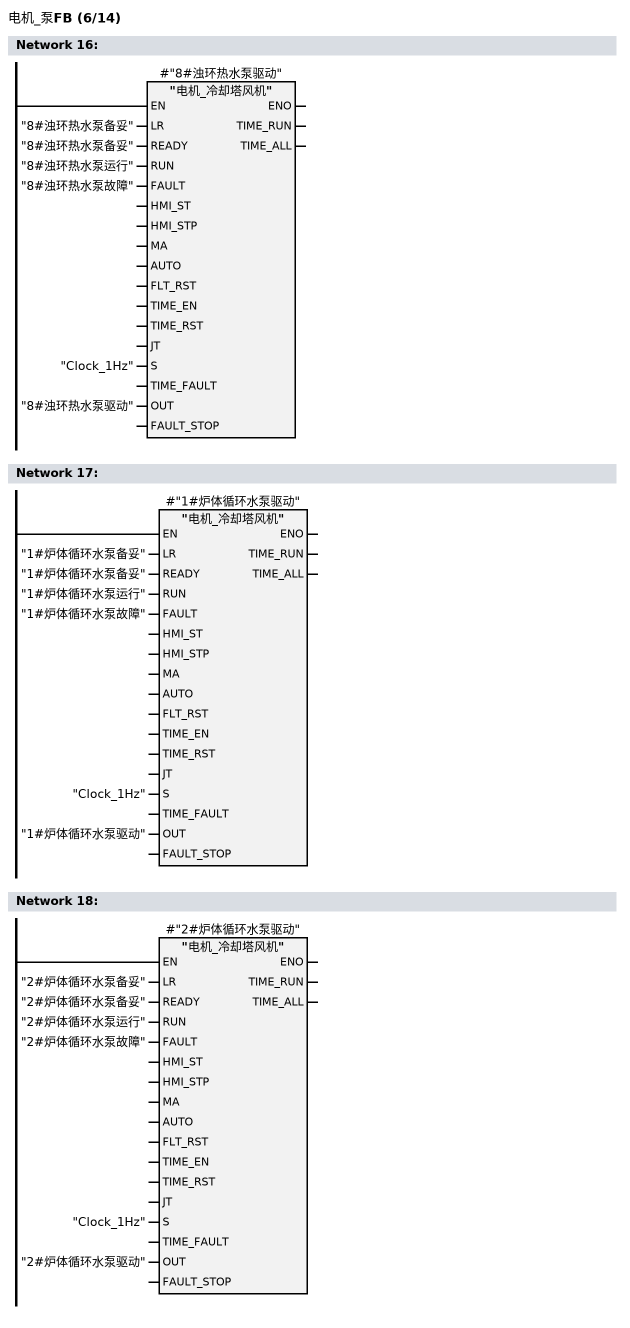
   RUNG wire#powerrail
      #"8#浊环热水泵驱动"(LR := "8#浊环热水泵备妥", READY := "8#浊环热水泵备妥", RUN := "8#浊环热水泵运行", FAULT := "8#浊环热水泵故障", HMI_ST :=, HMI_STP :=, MA :=, AUTO :=, FLT_RST :=, TIME_EN :=, TIME_RST :=, JT :=, S := "Clock_1Hz", TIME_FAULT :=, OUT := "8#浊环热水泵驱动", FAULT_STOP :=, TIME_RUN =>, TIME_ALL =>)
   END_RUNG
   // the same network as SCL:
   #"8#浊环热水泵驱动"(LR := "8#浊环热水泵备妥",   // "电机_冷却塔风机"
                READY := "8#浊环热水泵备妥",
                RUN := "8#浊环热水泵运行",
                FAULT := "8#浊环热水泵故障",
                S := "Clock_1Hz",
                OUT := "8#浊环热水泵驱动");
END_REGION

REGION Network 17
   RUNG wire#powerrail
      #"1#炉体循环水泵驱动"(LR := "1#炉体循环水泵备妥", READY := "1#炉体循环水泵备妥", RUN := "1#炉体循环水泵运行", FAULT := "1#炉体循环水泵故障", HMI_ST :=, HMI_STP :=, MA :=, AUTO :=, FLT_RST :=, TIME_EN :=, TIME_RST :=, JT :=, S := "Clock_1Hz", TIME_FAULT :=, OUT := "1#炉体循环水泵驱动", FAULT_STOP :=, TIME_RUN =>, TIME_ALL =>)
   END_RUNG
   // the same network as SCL:
   #"1#炉体循环水泵驱动"(LR := "1#炉体循环水泵备妥",   // "电机_冷却塔风机"
                 READY := "1#炉体循环水泵备妥",
                 RUN := "1#炉体循环水泵运行",
                 FAULT := "1#炉体循环水泵故障",
                 S := "Clock_1Hz",
                 OUT := "1#炉体循环水泵驱动");
END_REGION

REGION Network 18
   RUNG wire#powerrail
      #"2#炉体循环水泵驱动"(LR := "2#炉体循环水泵备妥", READY := "2#炉体循环水泵备妥", RUN := "2#炉体循环水泵运行", FAULT := "2#炉体循环水泵故障", HMI_ST :=, HMI_STP :=, MA :=, AUTO :=, FLT_RST :=, TIME_EN :=, TIME_RST :=, JT :=, S := "Clock_1Hz", TIME_FAULT :=, OUT := "2#炉体循环水泵驱动", FAULT_STOP :=, TIME_RUN =>, TIME_ALL =>)
   END_RUNG
   // the same network as SCL:
   #"2#炉体循环水泵驱动"(LR := "2#炉体循环水泵备妥",   // "电机_冷却塔风机"
                 READY := "2#炉体循环水泵备妥",
                 RUN := "2#炉体循环水泵运行",
                 FAULT := "2#炉体循环水泵故障",
                 S := "Clock_1Hz",
                 OUT := "2#炉体循环水泵驱动");
END_REGION

REGION Network 19
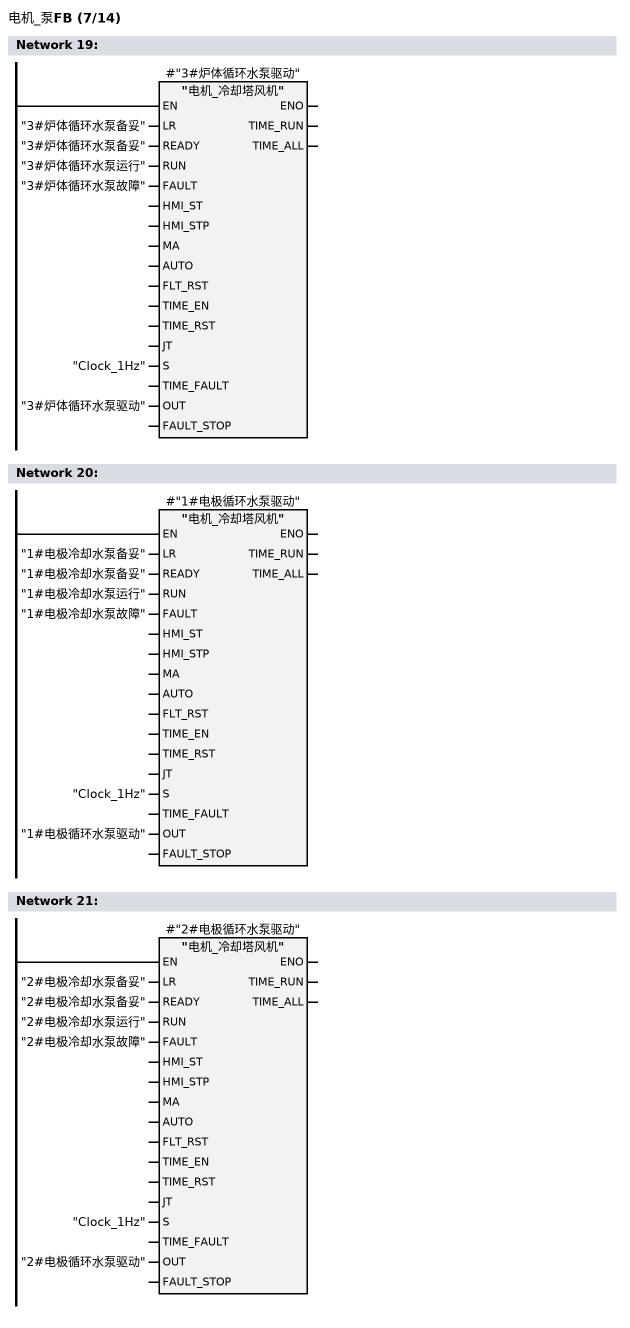
   RUNG wire#powerrail
      #"3#炉体循环水泵驱动"(LR := "3#炉体循环水泵备妥", READY := "3#炉体循环水泵备妥", RUN := "3#炉体循环水泵运行", FAULT := "3#炉体循环水泵故障", HMI_ST :=, HMI_STP :=, MA :=, AUTO :=, FLT_RST :=, TIME_EN :=, TIME_RST :=, JT :=, S := "Clock_1Hz", TIME_FAULT :=, OUT := "3#炉体循环水泵驱动", FAULT_STOP :=, TIME_RUN =>, TIME_ALL =>)
   END_RUNG
   // the same network as SCL:
   #"3#炉体循环水泵驱动"(LR := "3#炉体循环水泵备妥",   // "电机_冷却塔风机"
                 READY := "3#炉体循环水泵备妥",
                 RUN := "3#炉体循环水泵运行",
                 FAULT := "3#炉体循环水泵故障",
                 S := "Clock_1Hz",
                 OUT := "3#炉体循环水泵驱动");
END_REGION

REGION Network 20
   RUNG wire#powerrail
      #"1#电极循环水泵驱动"(LR := "1#电极冷却水泵备妥", READY := "1#电极冷却水泵备妥", RUN := "1#电极冷却水泵运行", FAULT := "1#电极冷却水泵故障", HMI_ST :=, HMI_STP :=, MA :=, AUTO :=, FLT_RST :=, TIME_EN :=, TIME_RST :=, JT :=, S := "Clock_1Hz", TIME_FAULT :=, OUT := "1#电极循环水泵驱动", FAULT_STOP :=, TIME_RUN =>, TIME_ALL =>)
   END_RUNG
   // the same network as SCL:
   #"1#电极循环水泵驱动"(LR := "1#电极冷却水泵备妥",   // "电机_冷却塔风机"
                 READY := "1#电极冷却水泵备妥",
                 RUN := "1#电极冷却水泵运行",
                 FAULT := "1#电极冷却水泵故障",
                 S := "Clock_1Hz",
                 OUT := "1#电极循环水泵驱动");
END_REGION

REGION Network 21
   RUNG wire#powerrail
      #"2#电极循环水泵驱动"(LR := "2#电极冷却水泵备妥", READY := "2#电极冷却水泵备妥", RUN := "2#电极冷却水泵运行", FAULT := "2#电极冷却水泵故障", HMI_ST :=, HMI_STP :=, MA :=, AUTO :=, FLT_RST :=, TIME_EN :=, TIME_RST :=, JT :=, S := "Clock_1Hz", TIME_FAULT :=, OUT := "2#电极循环水泵驱动", FAULT_STOP :=, TIME_RUN =>, TIME_ALL =>)
   END_RUNG
   // the same network as SCL:
   #"2#电极循环水泵驱动"(LR := "2#电极冷却水泵备妥",   // "电机_冷却塔风机"
                 READY := "2#电极冷却水泵备妥",
                 RUN := "2#电极冷却水泵运行",
                 FAULT := "2#电极冷却水泵故障",
                 S := "Clock_1Hz",
                 OUT := "2#电极循环水泵驱动");
END_REGION

REGION Network 22
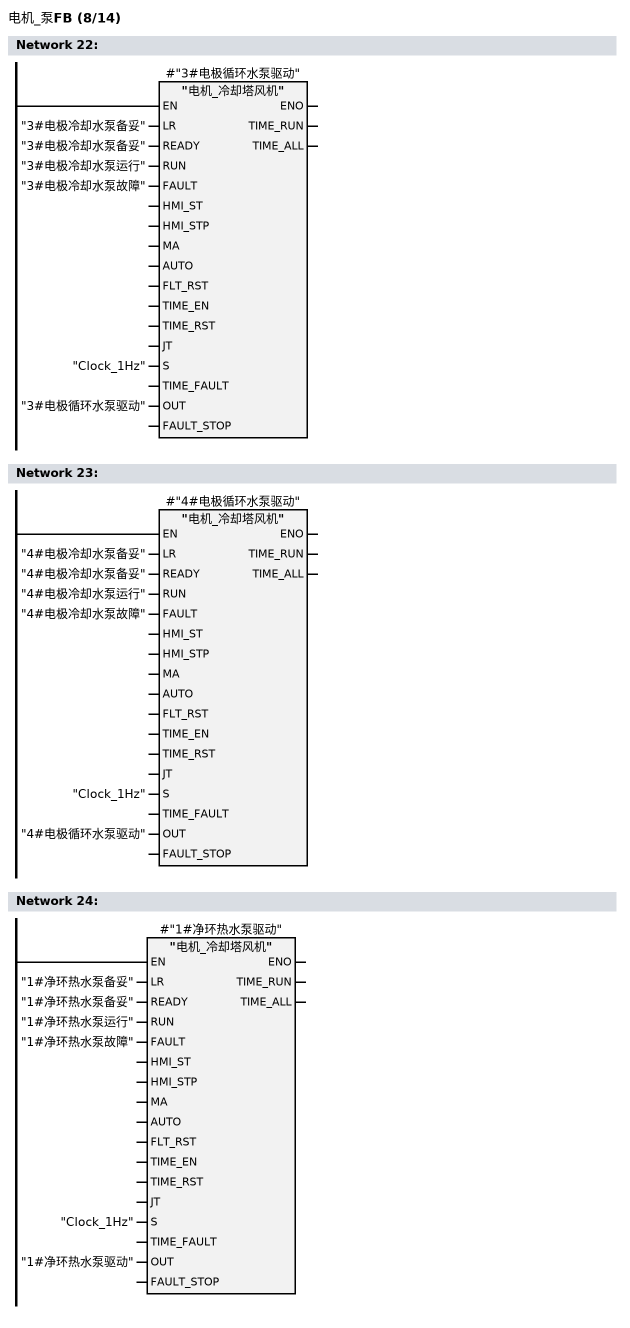
   RUNG wire#powerrail
      #"3#电极循环水泵驱动"(LR := "3#电极冷却水泵备妥", READY := "3#电极冷却水泵备妥", RUN := "3#电极冷却水泵运行", FAULT := "3#电极冷却水泵故障", HMI_ST :=, HMI_STP :=, MA :=, AUTO :=, FLT_RST :=, TIME_EN :=, TIME_RST :=, JT :=, S := "Clock_1Hz", TIME_FAULT :=, OUT := "3#电极循环水泵驱动", FAULT_STOP :=, TIME_RUN =>, TIME_ALL =>)
   END_RUNG
   // the same network as SCL:
   #"3#电极循环水泵驱动"(LR := "3#电极冷却水泵备妥",   // "电机_冷却塔风机"
                 READY := "3#电极冷却水泵备妥",
                 RUN := "3#电极冷却水泵运行",
                 FAULT := "3#电极冷却水泵故障",
                 S := "Clock_1Hz",
                 OUT := "3#电极循环水泵驱动");
END_REGION

REGION Network 23
   RUNG wire#powerrail
      #"4#电极循环水泵驱动"(LR := "4#电极冷却水泵备妥", READY := "4#电极冷却水泵备妥", RUN := "4#电极冷却水泵运行", FAULT := "4#电极冷却水泵故障", HMI_ST :=, HMI_STP :=, MA :=, AUTO :=, FLT_RST :=, TIME_EN :=, TIME_RST :=, JT :=, S := "Clock_1Hz", TIME_FAULT :=, OUT := "4#电极循环水泵驱动", FAULT_STOP :=, TIME_RUN =>, TIME_ALL =>)
   END_RUNG
   // the same network as SCL:
   #"4#电极循环水泵驱动"(LR := "4#电极冷却水泵备妥",   // "电机_冷却塔风机"
                 READY := "4#电极冷却水泵备妥",
                 RUN := "4#电极冷却水泵运行",
                 FAULT := "4#电极冷却水泵故障",
                 S := "Clock_1Hz",
                 OUT := "4#电极循环水泵驱动");
END_REGION

REGION Network 24
   RUNG wire#powerrail
      #"1#净环热水泵驱动"(LR := "1#净环热水泵备妥", READY := "1#净环热水泵备妥", RUN := "1#净环热水泵运行", FAULT := "1#净环热水泵故障", HMI_ST :=, HMI_STP :=, MA :=, AUTO :=, FLT_RST :=, TIME_EN :=, TIME_RST :=, JT :=, S := "Clock_1Hz", TIME_FAULT :=, OUT := "1#净环热水泵驱动", FAULT_STOP :=, TIME_RUN =>, TIME_ALL =>)
   END_RUNG
   // the same network as SCL:
   #"1#净环热水泵驱动"(LR := "1#净环热水泵备妥",   // "电机_冷却塔风机"
                READY := "1#净环热水泵备妥",
                RUN := "1#净环热水泵运行",
                FAULT := "1#净环热水泵故障",
                S := "Clock_1Hz",
                OUT := "1#净环热水泵驱动");
END_REGION

REGION Network 25
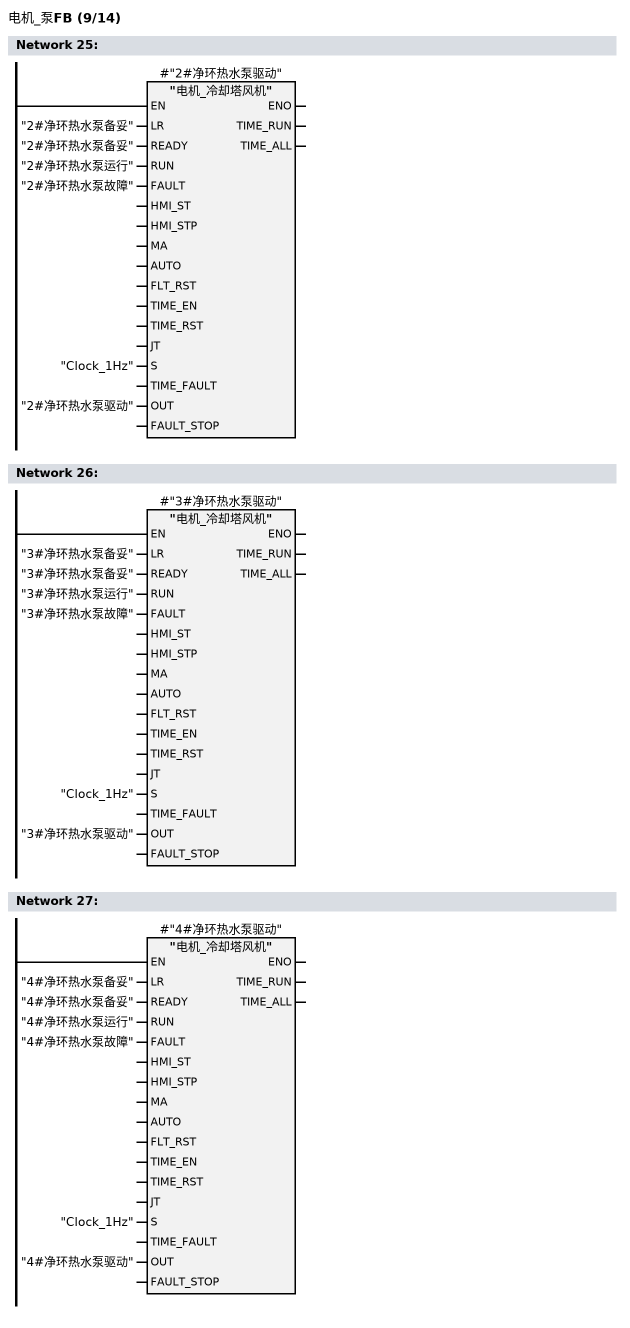
   RUNG wire#powerrail
      #"2#净环热水泵驱动"(LR := "2#净环热水泵备妥", READY := "2#净环热水泵备妥", RUN := "2#净环热水泵运行", FAULT := "2#净环热水泵故障", HMI_ST :=, HMI_STP :=, MA :=, AUTO :=, FLT_RST :=, TIME_EN :=, TIME_RST :=, JT :=, S := "Clock_1Hz", TIME_FAULT :=, OUT := "2#净环热水泵驱动", FAULT_STOP :=, TIME_RUN =>, TIME_ALL =>)
   END_RUNG
   // the same network as SCL:
   #"2#净环热水泵驱动"(LR := "2#净环热水泵备妥",   // "电机_冷却塔风机"
                READY := "2#净环热水泵备妥",
                RUN := "2#净环热水泵运行",
                FAULT := "2#净环热水泵故障",
                S := "Clock_1Hz",
                OUT := "2#净环热水泵驱动");
END_REGION

REGION Network 26
   RUNG wire#powerrail
      #"3#净环热水泵驱动"(LR := "3#净环热水泵备妥", READY := "3#净环热水泵备妥", RUN := "3#净环热水泵运行", FAULT := "3#净环热水泵故障", HMI_ST :=, HMI_STP :=, MA :=, AUTO :=, FLT_RST :=, TIME_EN :=, TIME_RST :=, JT :=, S := "Clock_1Hz", TIME_FAULT :=, OUT := "3#净环热水泵驱动", FAULT_STOP :=, TIME_RUN =>, TIME_ALL =>)
   END_RUNG
   // the same network as SCL:
   #"3#净环热水泵驱动"(LR := "3#净环热水泵备妥",   // "电机_冷却塔风机"
                READY := "3#净环热水泵备妥",
                RUN := "3#净环热水泵运行",
                FAULT := "3#净环热水泵故障",
                S := "Clock_1Hz",
                OUT := "3#净环热水泵驱动");
END_REGION

REGION Network 27
   RUNG wire#powerrail
      #"4#净环热水泵驱动"(LR := "4#净环热水泵备妥", READY := "4#净环热水泵备妥", RUN := "4#净环热水泵运行", FAULT := "4#净环热水泵故障", HMI_ST :=, HMI_STP :=, MA :=, AUTO :=, FLT_RST :=, TIME_EN :=, TIME_RST :=, JT :=, S := "Clock_1Hz", TIME_FAULT :=, OUT := "4#净环热水泵驱动", FAULT_STOP :=, TIME_RUN =>, TIME_ALL =>)
   END_RUNG
   // the same network as SCL:
   #"4#净环热水泵驱动"(LR := "4#净环热水泵备妥",   // "电机_冷却塔风机"
                READY := "4#净环热水泵备妥",
                RUN := "4#净环热水泵运行",
                FAULT := "4#净环热水泵故障",
                S := "Clock_1Hz",
                OUT := "4#净环热水泵驱动");
END_REGION

REGION Network 28
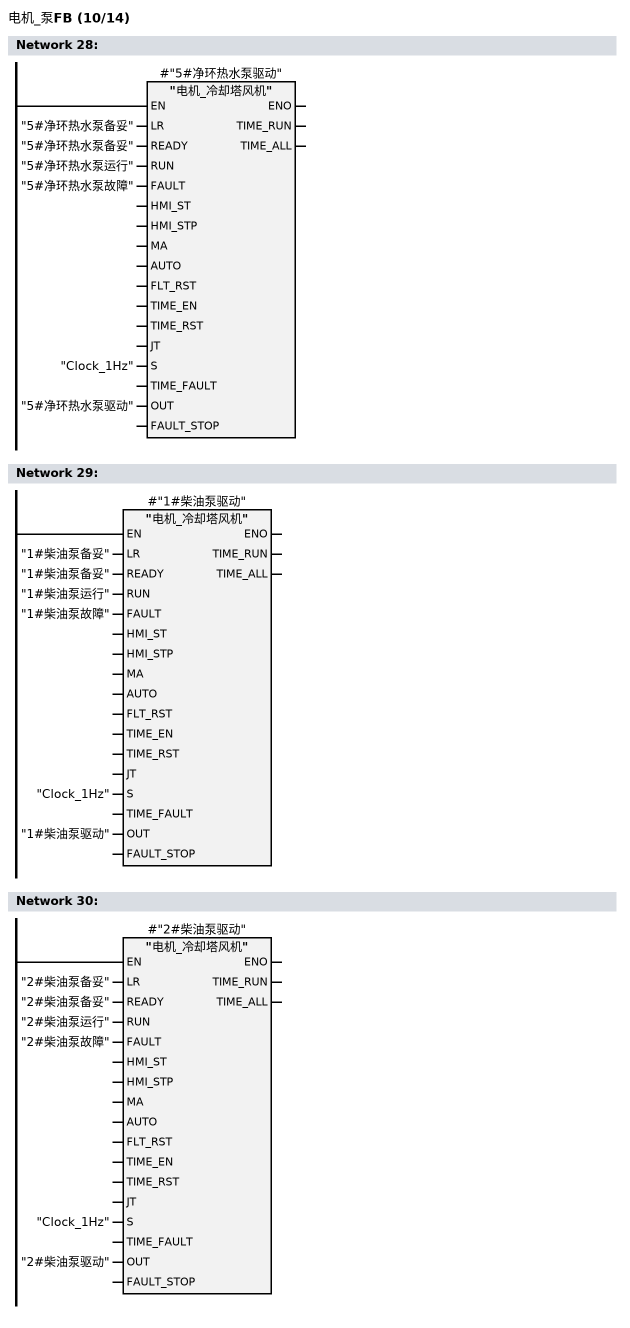
   RUNG wire#powerrail
      #"5#净环热水泵驱动"(LR := "5#净环热水泵备妥", READY := "5#净环热水泵备妥", RUN := "5#净环热水泵运行", FAULT := "5#净环热水泵故障", HMI_ST :=, HMI_STP :=, MA :=, AUTO :=, FLT_RST :=, TIME_EN :=, TIME_RST :=, JT :=, S := "Clock_1Hz", TIME_FAULT :=, OUT := "5#净环热水泵驱动", FAULT_STOP :=, TIME_RUN =>, TIME_ALL =>)
   END_RUNG
   // the same network as SCL:
   #"5#净环热水泵驱动"(LR := "5#净环热水泵备妥",   // "电机_冷却塔风机"
                READY := "5#净环热水泵备妥",
                RUN := "5#净环热水泵运行",
                FAULT := "5#净环热水泵故障",
                S := "Clock_1Hz",
                OUT := "5#净环热水泵驱动");
END_REGION

REGION Network 29
   RUNG wire#powerrail
      #"1#柴油泵驱动"(LR := "1#柴油泵备妥", READY := "1#柴油泵备妥", RUN := "1#柴油泵运行", FAULT := "1#柴油泵故障", HMI_ST :=, HMI_STP :=, MA :=, AUTO :=, FLT_RST :=, TIME_EN :=, TIME_RST :=, JT :=, S := "Clock_1Hz", TIME_FAULT :=, OUT := "1#柴油泵驱动", FAULT_STOP :=, TIME_RUN =>, TIME_ALL =>)
   END_RUNG
   // the same network as SCL:
   #"1#柴油泵驱动"(LR := "1#柴油泵备妥",   // "电机_冷却塔风机"
              READY := "1#柴油泵备妥",
              RUN := "1#柴油泵运行",
              FAULT := "1#柴油泵故障",
              S := "Clock_1Hz",
              OUT := "1#柴油泵驱动");
END_REGION

REGION Network 30
   RUNG wire#powerrail
      #"2#柴油泵驱动"(LR := "2#柴油泵备妥", READY := "2#柴油泵备妥", RUN := "2#柴油泵运行", FAULT := "2#柴油泵故障", HMI_ST :=, HMI_STP :=, MA :=, AUTO :=, FLT_RST :=, TIME_EN :=, TIME_RST :=, JT :=, S := "Clock_1Hz", TIME_FAULT :=, OUT := "2#柴油泵驱动", FAULT_STOP :=, TIME_RUN =>, TIME_ALL =>)
   END_RUNG
   // the same network as SCL:
   #"2#柴油泵驱动"(LR := "2#柴油泵备妥",   // "电机_冷却塔风机"
              READY := "2#柴油泵备妥",
              RUN := "2#柴油泵运行",
              FAULT := "2#柴油泵故障",
              S := "Clock_1Hz",
              OUT := "2#柴油泵驱动");
END_REGION

REGION Network 31
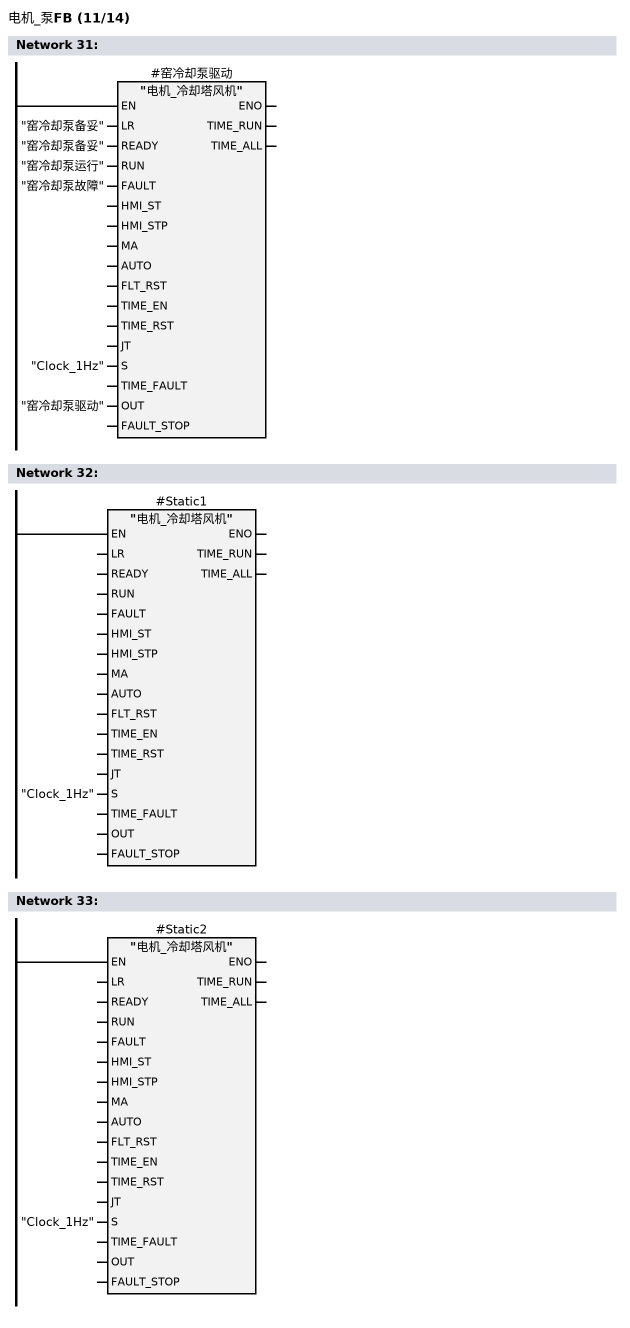
   RUNG wire#powerrail
      #窑冷却泵驱动(LR := "窑冷却泵备妥", READY := "窑冷却泵备妥", RUN := "窑冷却泵运行", FAULT := "窑冷却泵故障", HMI_ST :=, HMI_STP :=, MA :=, AUTO :=, FLT_RST :=, TIME_EN :=, TIME_RST :=, JT :=, S := "Clock_1Hz", TIME_FAULT :=, OUT := "窑冷却泵驱动", FAULT_STOP :=, TIME_RUN =>, TIME_ALL =>)
   END_RUNG
   // the same network as SCL:
   #窑冷却泵驱动(LR := "窑冷却泵备妥",   // "电机_冷却塔风机"
           READY := "窑冷却泵备妥",
           RUN := "窑冷却泵运行",
           FAULT := "窑冷却泵故障",
           S := "Clock_1Hz",
           OUT := "窑冷却泵驱动");
END_REGION

REGION Network 32
   RUNG wire#powerrail
      #Static1(LR :=, READY :=, RUN :=, FAULT :=, HMI_ST :=, HMI_STP :=, MA :=, AUTO :=, FLT_RST :=, TIME_EN :=, TIME_RST :=, JT :=, S := "Clock_1Hz", TIME_FAULT :=, OUT :=, FAULT_STOP :=, TIME_RUN =>, TIME_ALL =>)
   END_RUNG
   // the same network as SCL:
   #Static1(S := "Clock_1Hz");   // "电机_冷却塔风机"
END_REGION

REGION Network 33
   RUNG wire#powerrail
      #Static2(LR :=, READY :=, RUN :=, FAULT :=, HMI_ST :=, HMI_STP :=, MA :=, AUTO :=, FLT_RST :=, TIME_EN :=, TIME_RST :=, JT :=, S := "Clock_1Hz", TIME_FAULT :=, OUT :=, FAULT_STOP :=, TIME_RUN =>, TIME_ALL =>)
   END_RUNG
   // the same network as SCL:
   #Static2(S := "Clock_1Hz");   // "电机_冷却塔风机"
END_REGION

REGION Network 34
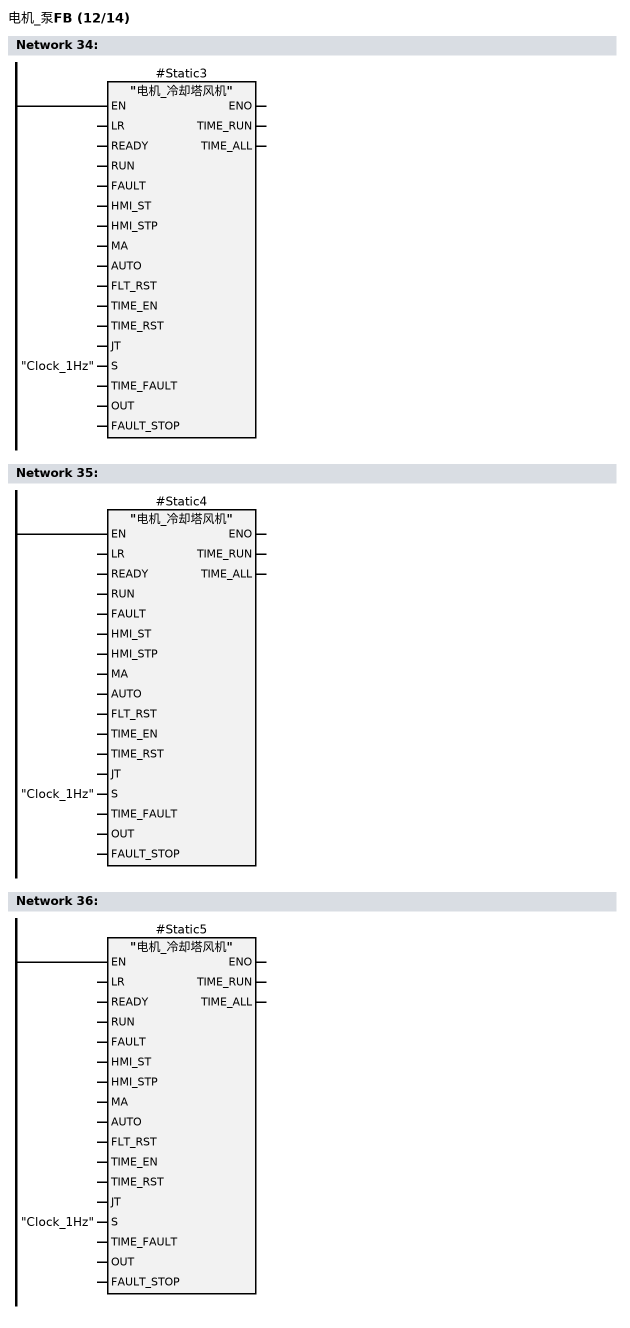
   RUNG wire#powerrail
      #Static3(LR :=, READY :=, RUN :=, FAULT :=, HMI_ST :=, HMI_STP :=, MA :=, AUTO :=, FLT_RST :=, TIME_EN :=, TIME_RST :=, JT :=, S := "Clock_1Hz", TIME_FAULT :=, OUT :=, FAULT_STOP :=, TIME_RUN =>, TIME_ALL =>)
   END_RUNG
   // the same network as SCL:
   #Static3(S := "Clock_1Hz");   // "电机_冷却塔风机"
END_REGION

REGION Network 35
   RUNG wire#powerrail
      #Static4(LR :=, READY :=, RUN :=, FAULT :=, HMI_ST :=, HMI_STP :=, MA :=, AUTO :=, FLT_RST :=, TIME_EN :=, TIME_RST :=, JT :=, S := "Clock_1Hz", TIME_FAULT :=, OUT :=, FAULT_STOP :=, TIME_RUN =>, TIME_ALL =>)
   END_RUNG
   // the same network as SCL:
   #Static4(S := "Clock_1Hz");   // "电机_冷却塔风机"
END_REGION

REGION Network 36
   RUNG wire#powerrail
      #Static5(LR :=, READY :=, RUN :=, FAULT :=, HMI_ST :=, HMI_STP :=, MA :=, AUTO :=, FLT_RST :=, TIME_EN :=, TIME_RST :=, JT :=, S := "Clock_1Hz", TIME_FAULT :=, OUT :=, FAULT_STOP :=, TIME_RUN =>, TIME_ALL =>)
   END_RUNG
   // the same network as SCL:
   #Static5(S := "Clock_1Hz");   // "电机_冷却塔风机"
END_REGION

REGION Network 37
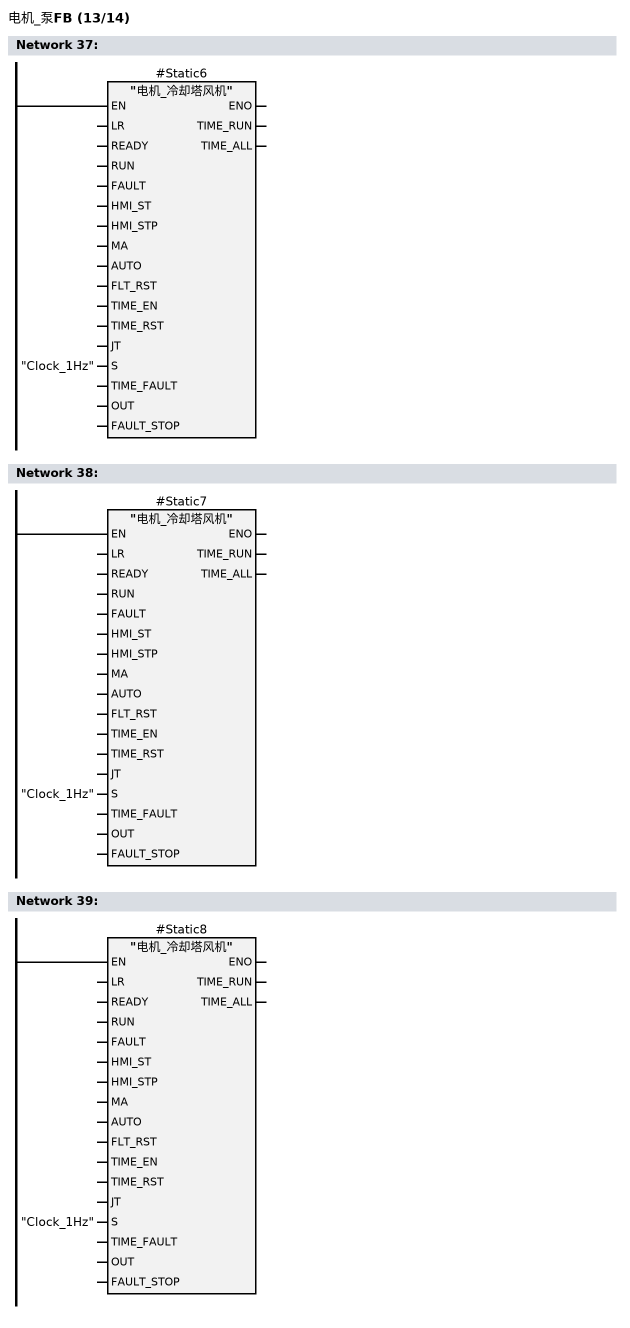
   RUNG wire#powerrail
      #Static6(LR :=, READY :=, RUN :=, FAULT :=, HMI_ST :=, HMI_STP :=, MA :=, AUTO :=, FLT_RST :=, TIME_EN :=, TIME_RST :=, JT :=, S := "Clock_1Hz", TIME_FAULT :=, OUT :=, FAULT_STOP :=, TIME_RUN =>, TIME_ALL =>)
   END_RUNG
   // the same network as SCL:
   #Static6(S := "Clock_1Hz");   // "电机_冷却塔风机"
END_REGION

REGION Network 38
   RUNG wire#powerrail
      #Static7(LR :=, READY :=, RUN :=, FAULT :=, HMI_ST :=, HMI_STP :=, MA :=, AUTO :=, FLT_RST :=, TIME_EN :=, TIME_RST :=, JT :=, S := "Clock_1Hz", TIME_FAULT :=, OUT :=, FAULT_STOP :=, TIME_RUN =>, TIME_ALL =>)
   END_RUNG
   // the same network as SCL:
   #Static7(S := "Clock_1Hz");   // "电机_冷却塔风机"
END_REGION

REGION Network 39
   RUNG wire#powerrail
      #Static8(LR :=, READY :=, RUN :=, FAULT :=, HMI_ST :=, HMI_STP :=, MA :=, AUTO :=, FLT_RST :=, TIME_EN :=, TIME_RST :=, JT :=, S := "Clock_1Hz", TIME_FAULT :=, OUT :=, FAULT_STOP :=, TIME_RUN =>, TIME_ALL =>)
   END_RUNG
   // the same network as SCL:
   #Static8(S := "Clock_1Hz");   // "电机_冷却塔风机"
END_REGION

REGION Network 40
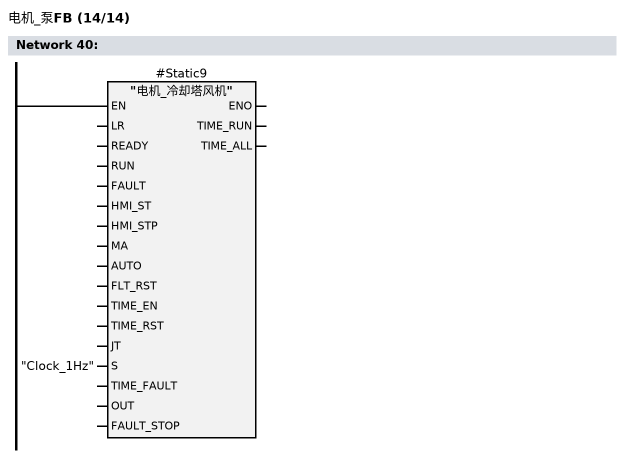
   RUNG wire#powerrail
      #Static9(LR :=, READY :=, RUN :=, FAULT :=, HMI_ST :=, HMI_STP :=, MA :=, AUTO :=, FLT_RST :=, TIME_EN :=, TIME_RST :=, JT :=, S := "Clock_1Hz", TIME_FAULT :=, OUT :=, FAULT_STOP :=, TIME_RUN =>, TIME_ALL =>)
   END_RUNG
   // the same network as SCL:
   #Static9(S := "Clock_1Hz");   // "电机_冷却塔风机"
END_REGION
END_FUNCTION_BLOCK

FUNCTION_BLOCK "FB14_DATA_ALARM"   // FB14, LAD
{ S7_Optimized_Access := 'FALSE' }
VERSION : 0.1
   VAR
      "PIW 256" : "FB330_DATA_ALARM";   // 1#炉体循环水泵管道压力
      "PIW 258" : "FB330_DATA_ALARM";   // 2#炉体循环水泵管道压力
      "PIW 260" : "FB330_DATA_ALARM";   // 3#炉体循环水泵管道压力
      "PIW 262" : "FB330_DATA_ALARM";   // 1#电极循环水泵管道压力
      "PIW 264" : "FB330_DATA_ALARM";   // 2#电极循环水泵管道压力
      "PIW 266" : "FB330_DATA_ALARM";   // 3#电极循环水泵管道压力
      "PIW 268" : "FB330_DATA_ALARM";   // 4#电极循环水泵管道压力
      "PIW 270" : "FB330_DATA_ALARM";   // 1#柴油泵管道压力
      "PIW 272" : "FB330_DATA_ALARM";   // 2#柴油泵管道压力
      "PIW 274" : "FB330_DATA_ALARM";   // 1#炉体循环水泵阀门开度
      "PIW 276" : "FB330_DATA_ALARM";   // 2#炉体循环水泵阀门开度
      "PIW 278" : "FB330_DATA_ALARM";   // 3#炉体循环水泵阀门开度
      "PIW 280" : "FB330_DATA_ALARM";   // 1#电极循环水泵阀门开度
      "PIW 282" : "FB330_DATA_ALARM";   // 2#电极循环水泵阀门开度
      "PIW 284" : "FB330_DATA_ALARM";   // 3#电极循环水泵阀门开度
      "PIW 286" : "FB330_DATA_ALARM";   // 4#电极循环水泵阀门开度
      "PIW 288" : "FB330_DATA_ALARM";   // 2#柴油泵阀门开度
      "PIW 290" : "FB330_DATA_ALARM";   // 1#净环热水管道压力
      "PIW 292" : "FB330_DATA_ALARM";   // 2#净环热水管道压力
      "PIW 294" : "FB330_DATA_ALARM";   // 3#净环热水管道压力
      "PIW 296" : "FB330_DATA_ALARM";   // 4#净环热水管道压力
      "PIW 298" : "FB330_DATA_ALARM";   // 5#净环热水管道压力
      "PIW 300" : "FB330_DATA_ALARM";   // 6#净环热水管道压力
      "PIW 302" : "FB330_DATA_ALARM";   // 1#净环热水阀门开度
      "PIW 304" : "FB330_DATA_ALARM";   // 2#净环热水阀门开度
      "PIW 306" : "FB330_DATA_ALARM";   // 3#净环热水阀门开度
      "PIW 308" : "FB330_DATA_ALARM";   // 4#净环热水阀门开度
      "PIW 310" : "FB330_DATA_ALARM";   // 5#净环热水阀门开度
      "PIW 312" : "FB330_DATA_ALARM";   // 6#净环热水阀门开度
      "PIW 314" : "FB330_DATA_ALARM";   // 1#外围补水阀门开度
      "PIW 316" : "FB330_DATA_ALARM";   // 2#外围补水阀门开度
      "PIW 318" : "FB330_DATA_ALARM";   // 1#水池液位
      "PIW 320" : "FB330_DATA_ALARM";   // 2#水池液位
      "PIW 322" : "FB330_DATA_ALARM";   // PIW322
      "PIW 324" : "FB330_DATA_ALARM";   // PIW324
      "PIW 326" : "FB330_DATA_ALARM";   // PIW326
      "PIW 328" : "FB330_DATA_ALARM";   // PIW328
      "PIW 330" : "FB330_DATA_ALARM";   // PIW330
      "PIW 332" : "FB330_DATA_ALARM";   // PIW332
      "PIW 334" : "FB330_DATA_ALARM";   // PIW334
      "PIW 336" : "FB330_DATA_ALARM";   // 1#浊环热水泵管道压力
      "PIW 338" : "FB330_DATA_ALARM";   // 2#浊环热水泵管道压力
      "PIW 340" : "FB330_DATA_ALARM";   // 3#浊环热水泵管道压力
      "PIW 342" : "FB330_DATA_ALARM";   // 4#浊环热水泵管道压力
      "PIW 344" : "FB330_DATA_ALARM";   // 5#浊环热水泵管道压力
      "PIW 346" : "FB330_DATA_ALARM";   // 6#浊环热水泵管道压力
      "PIW 348" : "FB330_DATA_ALARM";   // 7#浊环热水泵管道压力
      "PIW 350" : "FB330_DATA_ALARM";   // 8#浊环热水泵管道压力
      "PIW 352" : "FB330_DATA_ALARM";   // 1#冲渣热水阀门开度
      "PIW 354" : "FB330_DATA_ALARM";   // 2#冲渣热水阀门开度
      "PIW 356" : "FB330_DATA_ALARM";   // 3#冲渣热水阀门开度
      "PIW 358" : "FB330_DATA_ALARM";   // 4#冲渣热水阀门开度
      "PIW 360" : "FB330_DATA_ALARM";   // 5#冲渣热水阀门开度
      "PIW 362" : "FB330_DATA_ALARM";   // 6#冲渣热水阀门开度
      "PIW 364" : "FB330_DATA_ALARM";   // 7#冲渣热水阀门开度
      "PIW 366" : "FB330_DATA_ALARM";   // 8#冲渣热水阀门开度
      "PIW 368" : "FB330_DATA_ALARM";   // 1#冲渣泵管道压力
      "PIW 370" : "FB330_DATA_ALARM";   // 2#冲渣泵管道压力
      "PIW 372" : "FB330_DATA_ALARM";   // 3#冲渣泵管道压力
      "PIW 374" : "FB330_DATA_ALARM";   // 4#冲渣泵管道压力
      "PIW 376" : "FB330_DATA_ALARM";   // 5#冲渣泵管道压力
      "PIW 378" : "FB330_DATA_ALARM";   // 6#冲渣泵管道压力
      "PIW 380" : "FB330_DATA_ALARM";   // 7#冲渣泵管道压力
      "PIW 382" : "FB330_DATA_ALARM";   // 8#冲渣泵管道压力
      "PIW 384" : "FB330_DATA_ALARM";   // 1#冲渣阀门开度
      "PIW 386" : "FB330_DATA_ALARM";   // 2#冲渣阀门开度
      "PIW 388" : "FB330_DATA_ALARM";   // 3#冲渣阀门开度
      "PIW 390" : "FB330_DATA_ALARM";   // 4#冲渣阀门开度
      "PIW 392" : "FB330_DATA_ALARM";   // 5#冲渣阀门开度
      "PIW 394" : "FB330_DATA_ALARM";   // 6#冲渣阀门开度
      "PIW 396" : "FB330_DATA_ALARM";   // 7#冲渣阀门开度
      "PIW 398" : "FB330_DATA_ALARM";   // 8#冲渣阀门开度
      备用1 : "FB330_DATA_ALARM";
      备用2 : "FB330_DATA_ALARM";
      备用3 : "FB330_DATA_ALARM";
      备用4 : "FB330_DATA_ALARM";
      备用5 : "FB330_DATA_ALARM";
      备用6 : "FB330_DATA_ALARM";
      备用7 : "FB330_DATA_ALARM";
      备用8 : "FB330_DATA_ALARM";
   END_VAR
BEGIN

REGION Network 1
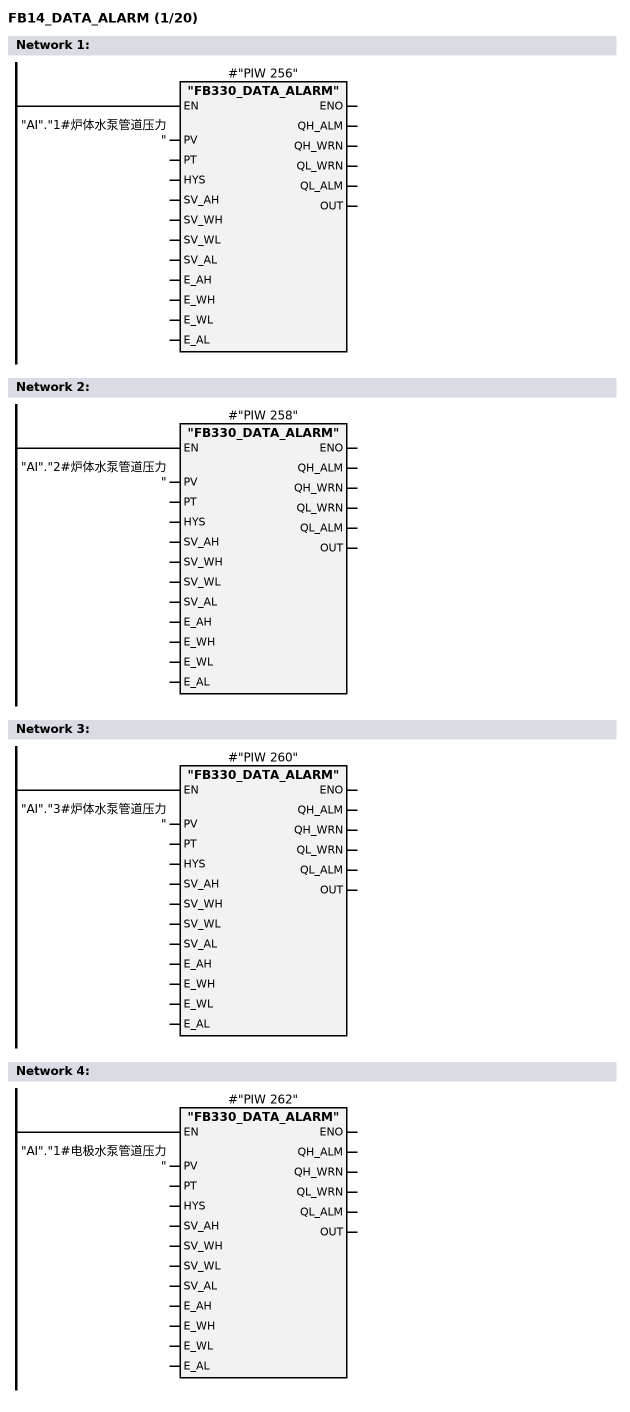
   RUNG wire#powerrail
      #"PIW 256"(PV := "AI"."1#炉体水泵管道压力", PT :=, HYS :=, SV_AH :=, SV_WH :=, SV_WL :=, SV_AL :=, E_AH :=, E_WH :=, E_WL :=, E_AL :=, QH_ALM =>, QH_WRN =>, QL_WRN =>, QL_ALM =>, OUT =>)
   END_RUNG
   // the same network as SCL:
   #"PIW 256"(PV := "AI"."1#炉体水泵管道压力");   // "FB330_DATA_ALARM"
END_REGION

REGION Network 2
   RUNG wire#powerrail
      #"PIW 258"(PV := "AI"."2#炉体水泵管道压力", PT :=, HYS :=, SV_AH :=, SV_WH :=, SV_WL :=, SV_AL :=, E_AH :=, E_WH :=, E_WL :=, E_AL :=, QH_ALM =>, QH_WRN =>, QL_WRN =>, QL_ALM =>, OUT =>)
   END_RUNG
   // the same network as SCL:
   #"PIW 258"(PV := "AI"."2#炉体水泵管道压力");   // "FB330_DATA_ALARM"
END_REGION

REGION Network 3
   RUNG wire#powerrail
      #"PIW 260"(PV := "AI"."3#炉体水泵管道压力", PT :=, HYS :=, SV_AH :=, SV_WH :=, SV_WL :=, SV_AL :=, E_AH :=, E_WH :=, E_WL :=, E_AL :=, QH_ALM =>, QH_WRN =>, QL_WRN =>, QL_ALM =>, OUT =>)
   END_RUNG
   // the same network as SCL:
   #"PIW 260"(PV := "AI"."3#炉体水泵管道压力");   // "FB330_DATA_ALARM"
END_REGION

REGION Network 4
   RUNG wire#powerrail
      #"PIW 262"(PV := "AI"."1#电极水泵管道压力", PT :=, HYS :=, SV_AH :=, SV_WH :=, SV_WL :=, SV_AL :=, E_AH :=, E_WH :=, E_WL :=, E_AL :=, QH_ALM =>, QH_WRN =>, QL_WRN =>, QL_ALM =>, OUT =>)
   END_RUNG
   // the same network as SCL:
   #"PIW 262"(PV := "AI"."1#电极水泵管道压力");   // "FB330_DATA_ALARM"
END_REGION

REGION Network 5
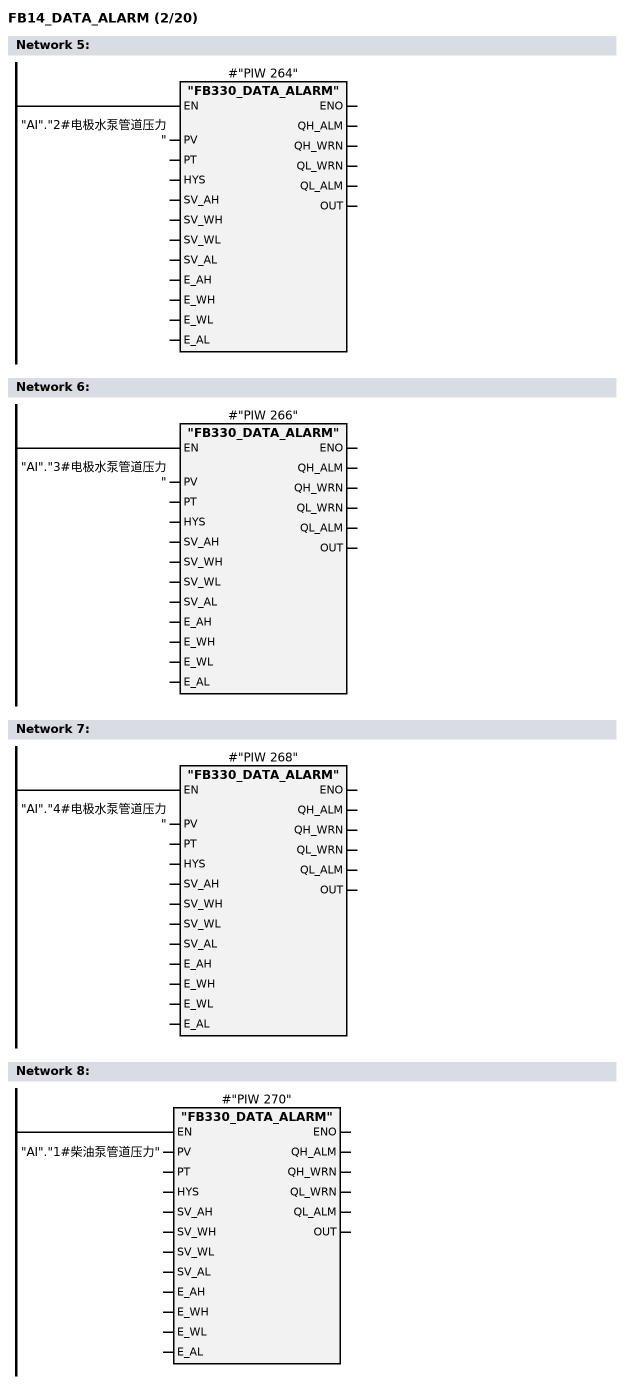
   RUNG wire#powerrail
      #"PIW 264"(PV := "AI"."2#电极水泵管道压力", PT :=, HYS :=, SV_AH :=, SV_WH :=, SV_WL :=, SV_AL :=, E_AH :=, E_WH :=, E_WL :=, E_AL :=, QH_ALM =>, QH_WRN =>, QL_WRN =>, QL_ALM =>, OUT =>)
   END_RUNG
   // the same network as SCL:
   #"PIW 264"(PV := "AI"."2#电极水泵管道压力");   // "FB330_DATA_ALARM"
END_REGION

REGION Network 6
   RUNG wire#powerrail
      #"PIW 266"(PV := "AI"."3#电极水泵管道压力", PT :=, HYS :=, SV_AH :=, SV_WH :=, SV_WL :=, SV_AL :=, E_AH :=, E_WH :=, E_WL :=, E_AL :=, QH_ALM =>, QH_WRN =>, QL_WRN =>, QL_ALM =>, OUT =>)
   END_RUNG
   // the same network as SCL:
   #"PIW 266"(PV := "AI"."3#电极水泵管道压力");   // "FB330_DATA_ALARM"
END_REGION

REGION Network 7
   RUNG wire#powerrail
      #"PIW 268"(PV := "AI"."4#电极水泵管道压力", PT :=, HYS :=, SV_AH :=, SV_WH :=, SV_WL :=, SV_AL :=, E_AH :=, E_WH :=, E_WL :=, E_AL :=, QH_ALM =>, QH_WRN =>, QL_WRN =>, QL_ALM =>, OUT =>)
   END_RUNG
   // the same network as SCL:
   #"PIW 268"(PV := "AI"."4#电极水泵管道压力");   // "FB330_DATA_ALARM"
END_REGION

REGION Network 8
   RUNG wire#powerrail
      #"PIW 270"(PV := "AI"."1#柴油泵管道压力", PT :=, HYS :=, SV_AH :=, SV_WH :=, SV_WL :=, SV_AL :=, E_AH :=, E_WH :=, E_WL :=, E_AL :=, QH_ALM =>, QH_WRN =>, QL_WRN =>, QL_ALM =>, OUT =>)
   END_RUNG
   // the same network as SCL:
   #"PIW 270"(PV := "AI"."1#柴油泵管道压力");   // "FB330_DATA_ALARM"
END_REGION

REGION Network 9